REGION Network 63: DeOx/ReOx Valave Configuration Done Sequence Delay
   // Get time value from HMI data
   RUNG wire#powerrail
      Move(in := "86_Times".VLV_CNFG_DN_DLY, out1 => "300_AUT_SEQ_TMRS_DB".VLV_CNFG_DN_DLY.PT)
   END_RUNG
   // the same network as SCL:
   "300_AUT_SEQ_TMRS_DB".VLV_CNFG_DN_DLY.PT := "86_Times".VLV_CNFG_DN_DLY;
END_REGION

REGION Network 64: Modify Maximum Step Time
   // To avoid time-out errors when value changed
   RUNG wire#powerrail
      Add(in1 := "300_AUT_SEQ_TMRS_DB".VLV_CNFG_DN_DLY.PT, in2 := T#100ms, out => "100_GCU_AUTO_SEQ_DB".STEP_410.MST)
   END_RUNG
   // the same network as SCL:
   "100_GCU_AUTO_SEQ_DB".STEP_410.MST := "300_AUT_SEQ_TMRS_DB".VLV_CNFG_DN_DLY.PT + T#100ms;
END_REGION

REGION Network 65: DeOx/ReOx Valave Configuration Done Sequence Delay
   // Run timer
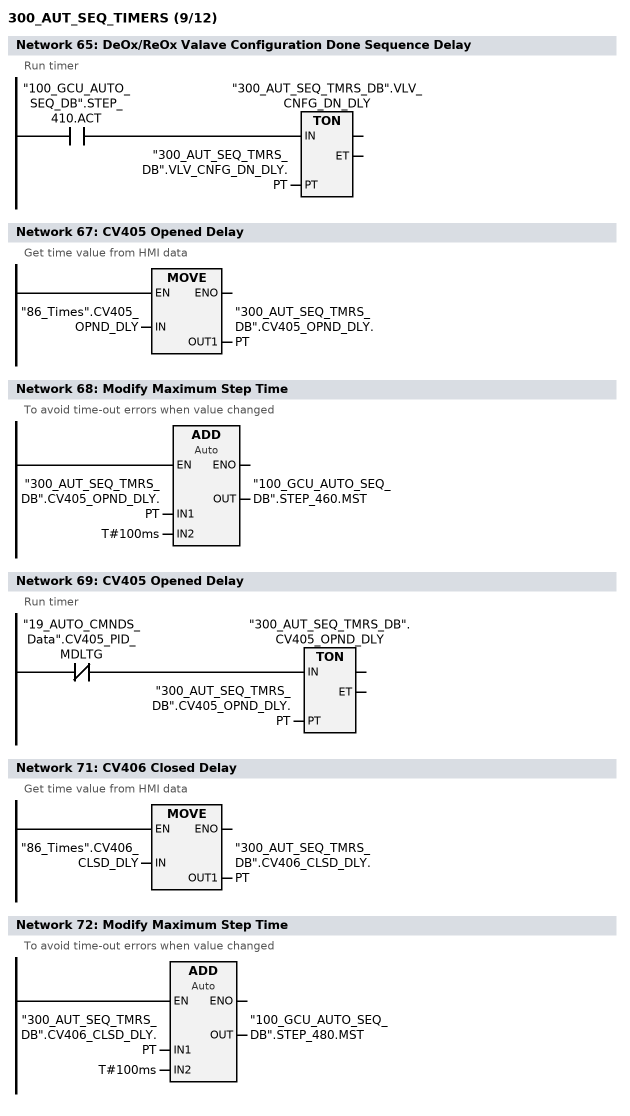
   "300_AUT_SEQ_TMRS_DB".VLV_CNFG_DN_DLY.TON(IN := "100_GCU_AUTO_SEQ_DB".STEP_410.ACT,
                           PT := "300_AUT_SEQ_TMRS_DB".VLV_CNFG_DN_DLY.PT);
END_REGION

REGION Network 67: CV405 Opened Delay
   // Get time value from HMI data
   RUNG wire#powerrail
      Move(in := "86_Times".CV405_OPND_DLY, out1 => "300_AUT_SEQ_TMRS_DB".CV405_OPND_DLY.PT)
   END_RUNG
   // the same network as SCL:
   "300_AUT_SEQ_TMRS_DB".CV405_OPND_DLY.PT := "86_Times".CV405_OPND_DLY;
END_REGION

REGION Network 68: Modify Maximum Step Time
   // To avoid time-out errors when value changed
   RUNG wire#powerrail
      Add(in1 := "300_AUT_SEQ_TMRS_DB".CV405_OPND_DLY.PT, in2 := T#100ms, out => "100_GCU_AUTO_SEQ_DB".STEP_460.MST)
   END_RUNG
   // the same network as SCL:
   "100_GCU_AUTO_SEQ_DB".STEP_460.MST := "300_AUT_SEQ_TMRS_DB".CV405_OPND_DLY.PT + T#100ms;
END_REGION

REGION Network 69: CV405 Opened Delay
   // Run timer
   "300_AUT_SEQ_TMRS_DB".CV405_OPND_DLY.TON(IN := NOT "19_AUTO_CMNDS_Data".CV405_PID_MDLTG,
                           PT := "300_AUT_SEQ_TMRS_DB".CV405_OPND_DLY.PT);
END_REGION

REGION Network 71: CV406 Closed Delay
   // Get time value from HMI data
   RUNG wire#powerrail
      Move(in := "86_Times".CV406_CLSD_DLY, out1 => "300_AUT_SEQ_TMRS_DB".CV406_CLSD_DLY.PT)
   END_RUNG
   // the same network as SCL:
   "300_AUT_SEQ_TMRS_DB".CV406_CLSD_DLY.PT := "86_Times".CV406_CLSD_DLY;
END_REGION

REGION Network 72: Modify Maximum Step Time
   // To avoid time-out errors when value changed
   RUNG wire#powerrail
      Add(in1 := "300_AUT_SEQ_TMRS_DB".CV406_CLSD_DLY.PT, in2 := T#100ms, out => "100_GCU_AUTO_SEQ_DB".STEP_480.MST)
   END_RUNG
   // the same network as SCL:
   "100_GCU_AUTO_SEQ_DB".STEP_480.MST := "300_AUT_SEQ_TMRS_DB".CV406_CLSD_DLY.PT + T#100ms;
END_REGION

REGION Network 73: CV406 Closed Delay
   // Run timer
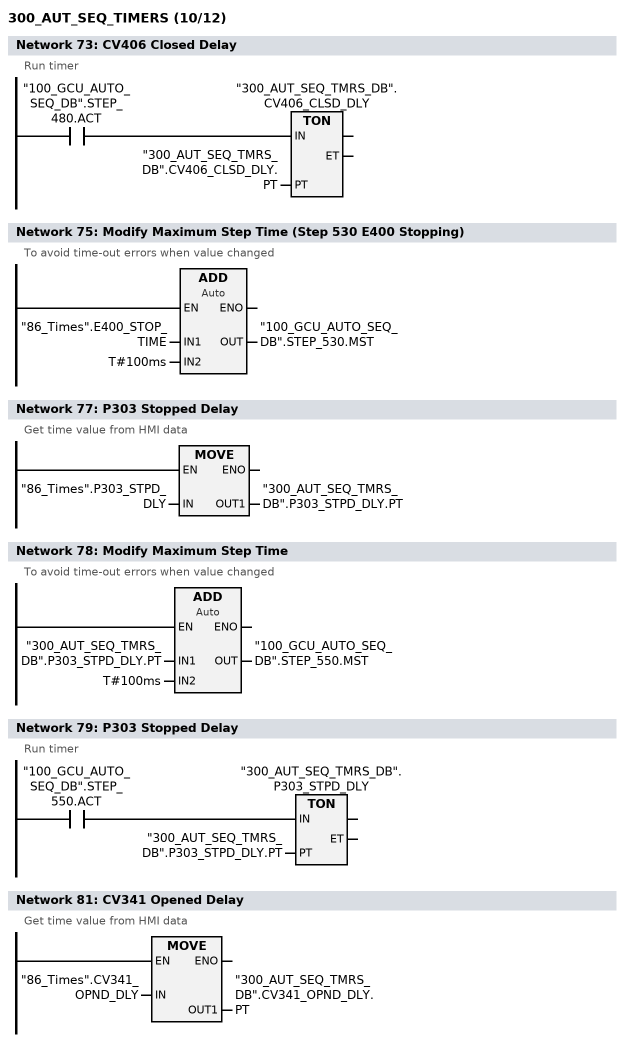
   "300_AUT_SEQ_TMRS_DB".CV406_CLSD_DLY.TON(IN := "100_GCU_AUTO_SEQ_DB".STEP_480.ACT,
                           PT := "300_AUT_SEQ_TMRS_DB".CV406_CLSD_DLY.PT);
END_REGION

REGION Network 75: Modify Maximum Step Time (Step 530 E400 Stopping)
   // To avoid time-out errors when value changed
   RUNG wire#powerrail
      Add(in1 := "86_Times".E400_STOP_TIME, in2 := T#100ms, out => "100_GCU_AUTO_SEQ_DB".STEP_530.MST)
   END_RUNG
   // the same network as SCL:
   "100_GCU_AUTO_SEQ_DB".STEP_530.MST := "86_Times".E400_STOP_TIME + T#100ms;
END_REGION

REGION Network 77: P303 Stopped Delay
   // Get time value from HMI data
   RUNG wire#powerrail
      Move(in := "86_Times".P303_STPD_DLY, out1 => "300_AUT_SEQ_TMRS_DB".P303_STPD_DLY.PT)
   END_RUNG
   // the same network as SCL:
   "300_AUT_SEQ_TMRS_DB".P303_STPD_DLY.PT := "86_Times".P303_STPD_DLY;
END_REGION

REGION Network 78: Modify Maximum Step Time
   // To avoid time-out errors when value changed
   RUNG wire#powerrail
      Add(in1 := "300_AUT_SEQ_TMRS_DB".P303_STPD_DLY.PT, in2 := T#100ms, out => "100_GCU_AUTO_SEQ_DB".STEP_550.MST)
   END_RUNG
   // the same network as SCL:
   "100_GCU_AUTO_SEQ_DB".STEP_550.MST := "300_AUT_SEQ_TMRS_DB".P303_STPD_DLY.PT + T#100ms;
END_REGION

REGION Network 79: P303 Stopped Delay
   // Run timer
   "300_AUT_SEQ_TMRS_DB".P303_STPD_DLY.TON(IN := "100_GCU_AUTO_SEQ_DB".STEP_550.ACT,
                           PT := "300_AUT_SEQ_TMRS_DB".P303_STPD_DLY.PT);
END_REGION

REGION Network 81: CV341 Opened Delay
   // Get time value from HMI data
   RUNG wire#powerrail
      Move(in := "86_Times".CV341_OPND_DLY, out1 => "300_AUT_SEQ_TMRS_DB".CV341_OPND_DLY.PT)
   END_RUNG
   // the same network as SCL:
   "300_AUT_SEQ_TMRS_DB".CV341_OPND_DLY.PT := "86_Times".CV341_OPND_DLY;
END_REGION

REGION Network 82: Modify Maximum Step Time
   // To avoid time-out errors when value changed
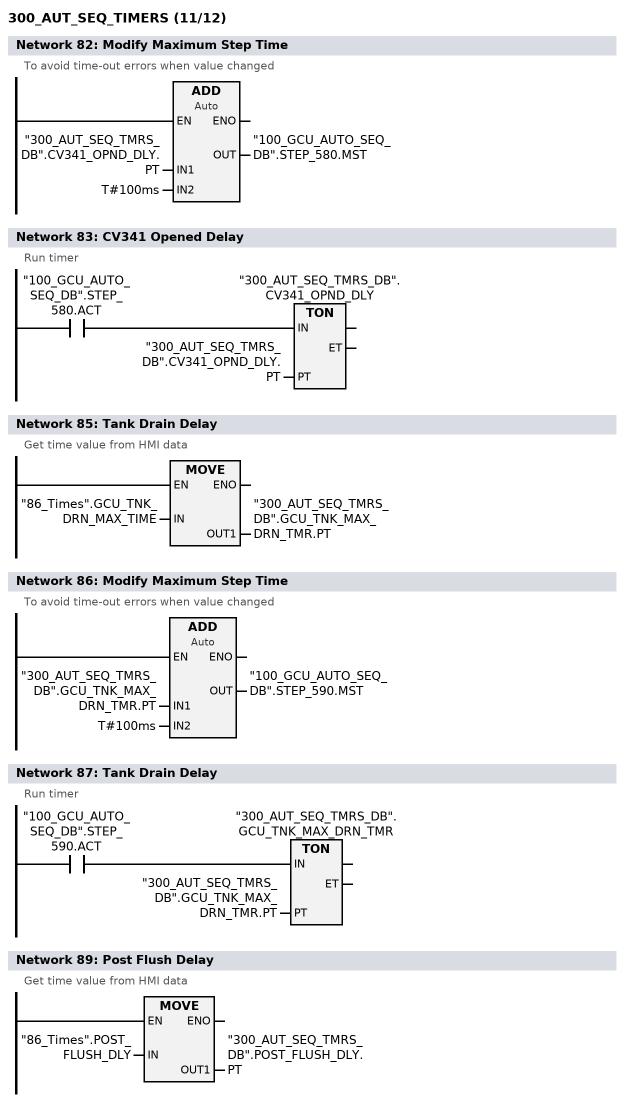
   RUNG wire#powerrail
      Add(in1 := "300_AUT_SEQ_TMRS_DB".CV341_OPND_DLY.PT, in2 := T#100ms, out => "100_GCU_AUTO_SEQ_DB".STEP_580.MST)
   END_RUNG
   // the same network as SCL:
   "100_GCU_AUTO_SEQ_DB".STEP_580.MST := "300_AUT_SEQ_TMRS_DB".CV341_OPND_DLY.PT + T#100ms;
END_REGION

REGION Network 83: CV341 Opened Delay
   // Run timer
   "300_AUT_SEQ_TMRS_DB".CV341_OPND_DLY.TON(IN := "100_GCU_AUTO_SEQ_DB".STEP_580.ACT,
                           PT := "300_AUT_SEQ_TMRS_DB".CV341_OPND_DLY.PT);
END_REGION

REGION Network 85: Tank Drain Delay
   // Get time value from HMI data
   RUNG wire#powerrail
      Move(in := "86_Times".GCU_TNK_DRN_MAX_TIME, out1 => "300_AUT_SEQ_TMRS_DB".GCU_TNK_MAX_DRN_TMR.PT)
   END_RUNG
   // the same network as SCL:
   "300_AUT_SEQ_TMRS_DB".GCU_TNK_MAX_DRN_TMR.PT := "86_Times".GCU_TNK_DRN_MAX_TIME;
END_REGION

REGION Network 86: Modify Maximum Step Time
   // To avoid time-out errors when value changed
   RUNG wire#powerrail
      Add(in1 := "300_AUT_SEQ_TMRS_DB".GCU_TNK_MAX_DRN_TMR.PT, in2 := T#100ms, out => "100_GCU_AUTO_SEQ_DB".STEP_590.MST)
   END_RUNG
   // the same network as SCL:
   "100_GCU_AUTO_SEQ_DB".STEP_590.MST := "300_AUT_SEQ_TMRS_DB".GCU_TNK_MAX_DRN_TMR.PT + T#100ms;
END_REGION

REGION Network 87: Tank Drain Delay
   // Run timer
   "300_AUT_SEQ_TMRS_DB".GCU_TNK_MAX_DRN_TMR.TON(IN := "100_GCU_AUTO_SEQ_DB".STEP_590.ACT,
                           PT := "300_AUT_SEQ_TMRS_DB".GCU_TNK_MAX_DRN_TMR.PT);
END_REGION

REGION Network 89: Post Flush Delay
   // Get time value from HMI data
   RUNG wire#powerrail
      Move(in := "86_Times".POST_FLUSH_DLY, out1 => "300_AUT_SEQ_TMRS_DB".POST_FLUSH_DLY.PT)
   END_RUNG
   // the same network as SCL:
   "300_AUT_SEQ_TMRS_DB".POST_FLUSH_DLY.PT := "86_Times".POST_FLUSH_DLY;
END_REGION

REGION Network 90: Modify Maximum Step Time
   // To avoid time-out errors when value changed
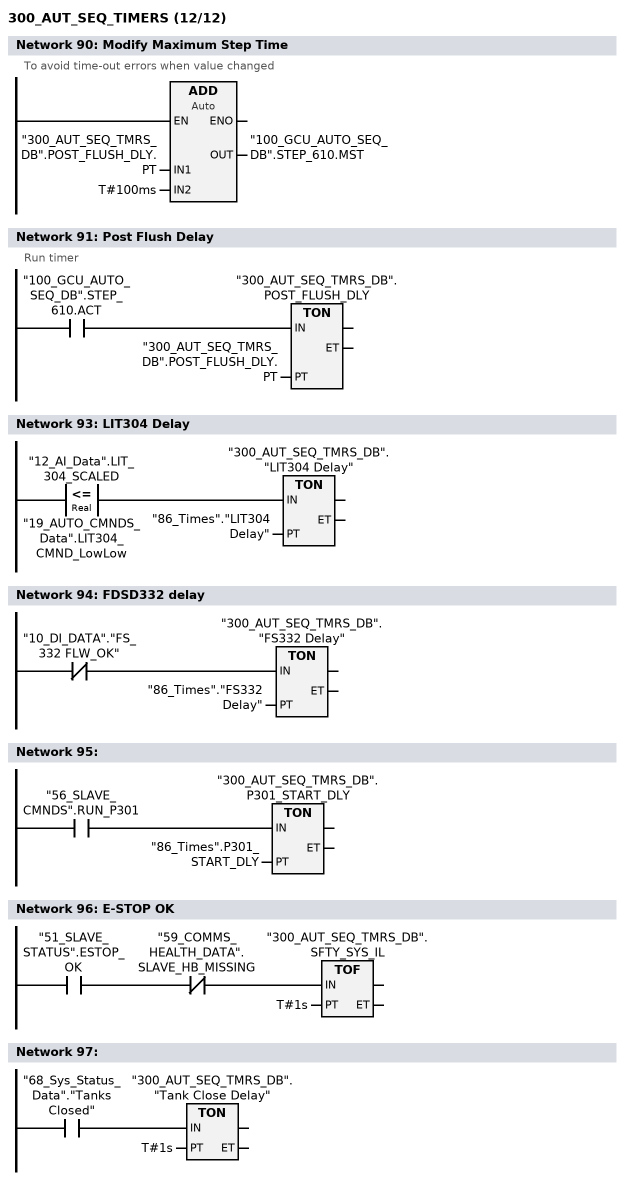
   RUNG wire#powerrail
      Add(in1 := "300_AUT_SEQ_TMRS_DB".POST_FLUSH_DLY.PT, in2 := T#100ms, out => "100_GCU_AUTO_SEQ_DB".STEP_610.MST)
   END_RUNG
   // the same network as SCL:
   "100_GCU_AUTO_SEQ_DB".STEP_610.MST := "300_AUT_SEQ_TMRS_DB".POST_FLUSH_DLY.PT + T#100ms;
END_REGION

REGION Network 91: Post Flush Delay
   // Run timer
   "300_AUT_SEQ_TMRS_DB".POST_FLUSH_DLY.TON(IN := "100_GCU_AUTO_SEQ_DB".STEP_610.ACT,
                           PT := "300_AUT_SEQ_TMRS_DB".POST_FLUSH_DLY.PT);
END_REGION

REGION Network 93: LIT304 Delay
   "300_AUT_SEQ_TMRS_DB"."LIT304 Delay".TON(IN := "12_AI_Data".LIT_304_SCALED <= "19_AUTO_CMNDS_Data".LIT304_CMND_LowLow,
                           PT := "86_Times"."LIT304 Delay");
END_REGION

REGION Network 94: FDSD332 delay
   "300_AUT_SEQ_TMRS_DB"."FS332 Delay".TON(IN := NOT "10_DI_DATA"."FS_332 FLW_OK",
                           PT := "86_Times"."FS332 Delay");
END_REGION

REGION Network 95
   "300_AUT_SEQ_TMRS_DB".P301_START_DLY.TON(IN := "56_SLAVE_CMNDS".RUN_P301, PT := "86_Times".P301_START_DLY);
END_REGION

REGION Network 96: E-STOP OK
   "300_AUT_SEQ_TMRS_DB".SFTY_SYS_IL.TOF(IN := "51_SLAVE_STATUS".ESTOP_OK AND NOT "59_COMMS_HEALTH_DATA".SLAVE_HB_MISSING,
                           PT := T#1s);
END_REGION

REGION Network 97
   "300_AUT_SEQ_TMRS_DB"."Tank Close Delay".TON(IN := "68_Sys_Status_Data"."Tanks Closed", PT := T#1s);
END_REGION
END_FUNCTION

// folder: 50 - 59 PLC Communication

FUNCTION "51_GET_SLAVE_DATA" : Void   // FC51, LAD
TITLE = Get Slave Status Data
{ S7_Optimized_Access := 'TRUE' }
AUTHOR : JRS
VERSION : 0.1
// Code for getting status data from the slave PLC (IGG)
   VAR_TEMP
      RET_VAL_1 : Int;
   END_VAR
BEGIN

REGION Network 1: Get Slave Status Data
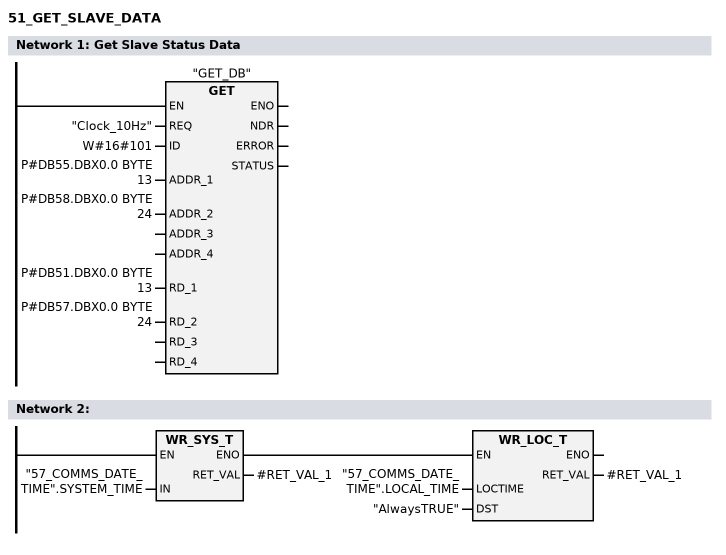
   "GET_DB"(REQ := "Clock_10Hz",   // GET
            ID := W#16#101,
            ADDR_1 := P#DB55.DBX0.0 BYTE 13,
            ADDR_2 := P#DB58.DBX0.0 BYTE 24,
            RD_1 := P#DB51.DBX0.0 BYTE 13,
            RD_2 := P#DB57.DBX0.0 BYTE 24);
END_REGION

REGION Network 2
   // ENO of a box is taken as its EN; it also drops when the box reports an error
   #RET_VAL_1 := WR_SYS_T(IN := "57_COMMS_DATE_TIME".SYSTEM_TIME);
   #RET_VAL_1 := WR_LOC_T(LOCTIME := "57_COMMS_DATE_TIME".LOCAL_TIME, DST := "AlwaysTRUE");
END_REGION
END_FUNCTION

FUNCTION "56_PUT_SLAVE_DATA" : Void   // FC56, LAD
TITLE = Put Slave Comands Data
{ S7_Optimized_Access := 'TRUE' }
AUTHOR : JRS
VERSION : 0.1
// Code for sending commands to the slave PLC (IGG)
BEGIN

REGION Network 1: PUT Slave Commands
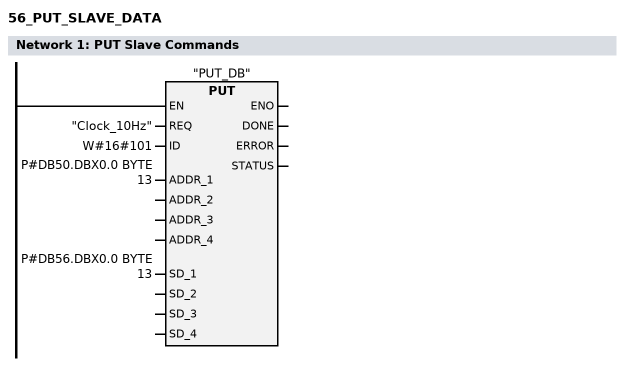
   "PUT_DB"(REQ := "Clock_10Hz", ID := W#16#101, ADDR_1 := P#DB50.DBX0.0 BYTE 13, SD_1 := P#DB56.DBX0.0 BYTE 13);   // PUT
END_REGION
END_FUNCTION

FUNCTION "59_COMMS_HEALTH" : Void   // FC59, LAD
TITLE = Communications Heart Beat
{ S7_Optimized_Access := 'TRUE' }
AUTHOR : JRS
VERSION : 0.1
// Code for communications heart beat bit
   VAR_TEMP   // added for the SCL form of the ladder/FBD networks
      _w1 : Bool;
   END_VAR
BEGIN

REGION Network 1: Local Heart Beat
   // Flip flop for status to other PLC's
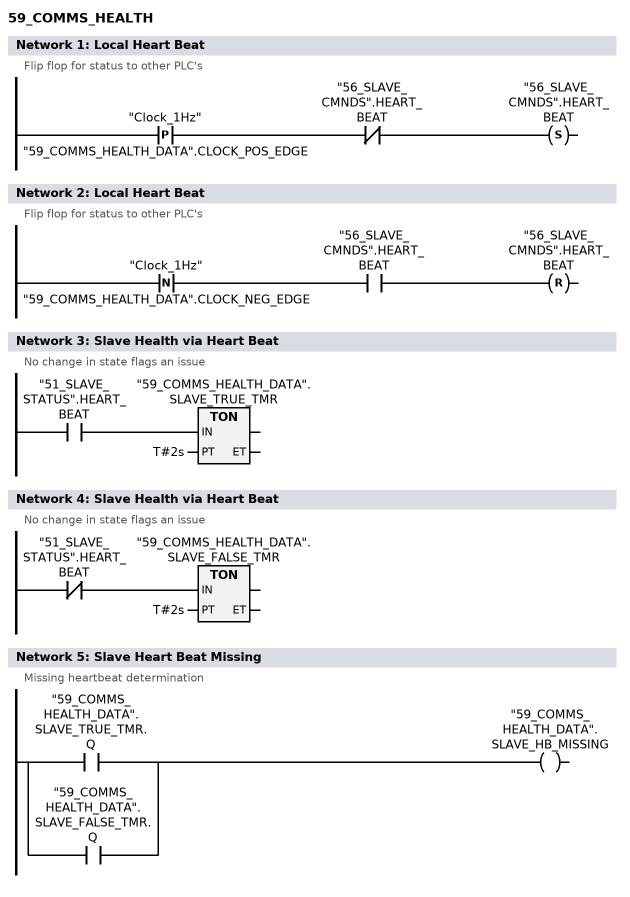
   RUNG wire#powerrail
      P_Contact(operand := "Clock_1Hz", bit := "59_COMMS_HEALTH_DATA".CLOCK_POS_EDGE)
      I_Contact( "56_SLAVE_CMNDS".HEART_BEAT )
      S_Coil( "56_SLAVE_CMNDS".HEART_BEAT )
   END_RUNG
   // the same network as SCL:
   #_w1 := "Clock_1Hz" AND NOT "59_COMMS_HEALTH_DATA".CLOCK_POS_EDGE;   // rising edge of "Clock_1Hz"
   "59_COMMS_HEALTH_DATA".CLOCK_POS_EDGE := "Clock_1Hz";
   IF #_w1 AND NOT "56_SLAVE_CMNDS".HEART_BEAT THEN "56_SLAVE_CMNDS".HEART_BEAT := TRUE; END_IF;
END_REGION

REGION Network 2: Local Heart Beat
   // Flip flop for status to other PLC's
   RUNG wire#powerrail
      N_Contact(operand := "Clock_1Hz", bit := "59_COMMS_HEALTH_DATA".CLOCK_NEG_EDGE)
      Contact( "56_SLAVE_CMNDS".HEART_BEAT )
      R_Coil( "56_SLAVE_CMNDS".HEART_BEAT )
   END_RUNG
   // the same network as SCL:
   #_w1 := NOT "Clock_1Hz" AND "59_COMMS_HEALTH_DATA".CLOCK_NEG_EDGE;   // falling edge of "Clock_1Hz"
   "59_COMMS_HEALTH_DATA".CLOCK_NEG_EDGE := "Clock_1Hz";
   IF #_w1 AND "56_SLAVE_CMNDS".HEART_BEAT THEN "56_SLAVE_CMNDS".HEART_BEAT := FALSE; END_IF;
END_REGION

REGION Network 3: Slave Health via Heart Beat
   // No change in state flags an issue
   "59_COMMS_HEALTH_DATA".SLAVE_TRUE_TMR.TON(IN := "51_SLAVE_STATUS".HEART_BEAT, PT := T#2s);
END_REGION

REGION Network 4: Slave Health via Heart Beat
   // No change in state flags an issue
   "59_COMMS_HEALTH_DATA".SLAVE_FALSE_TMR.TON(IN := NOT "51_SLAVE_STATUS".HEART_BEAT, PT := T#2s);
END_REGION

REGION Network 5: Slave Heart Beat Missing
   // Missing heartbeat determination
   RUNG wire#powerrail
      Contact( "59_COMMS_HEALTH_DATA".SLAVE_TRUE_TMR.Q )
      wire#w1
      Coil( "59_COMMS_HEALTH_DATA".SLAVE_HB_MISSING )
   END_RUNG
   RUNG wire#powerrail
      Contact( "59_COMMS_HEALTH_DATA".SLAVE_FALSE_TMR.Q )
   END_RUNG wire#w1
   // the same network as SCL:
   "59_COMMS_HEALTH_DATA".SLAVE_HB_MISSING := "59_COMMS_HEALTH_DATA".SLAVE_TRUE_TMR.Q OR "59_COMMS_HEALTH_DATA".SLAVE_FALSE_TMR.Q;
END_REGION
END_FUNCTION

// folder: 500 - 699 Standard FBs

FUNCTION_BLOCK "500_SEQ_STEP"   // FB500, LAD
{ S7_Optimized_Access := 'TRUE' }
VERSION : 0.1
   VAR_INPUT
      SN : Int;   // Step number
      CS : Int;   // Current step
      MST : Time;   // Maximum step time
      SC : Bool;   // Step complete
      BPFLT : Bool;   // Bypass fault
   END_VAR
   VAR_OUTPUT
      ACT : Bool;   // Active
      DN : Bool;   // Done
   END_VAR
   VAR_IN_OUT
      AMST : Time;   // Actual maximum step time
      FLT : Bool;   // Timed out
   END_VAR
   VAR
      RNG : Bool;   // Running
   END_VAR
   VAR RETAIN
      STP_MAX_TIM : TON_TIME;   // Maximum step time
   END_VAR
   VAR
      IEC_Timer_0_Instance : TOF_TIME;
   END_VAR
BEGIN

REGION Network 1: Step Active
   // When step number is active, it is also running
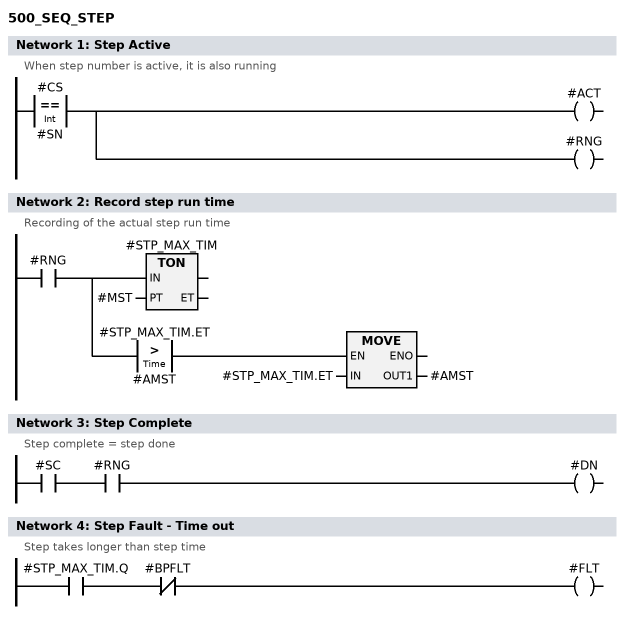
   RUNG wire#powerrail
      { S7_Templates := "SrcType := Int" } EQ_Contact(in1 := #CS, in2 := #SN)
      wire#w1
      Coil( #ACT )
   END_RUNG
   RUNG wire#w1
      Coil( #RNG )
   END_RUNG
   // the same network as SCL:
   #ACT := #CS = #SN;
   #RNG := #ACT;
END_REGION

REGION Network 2: Record step run time
   // Recording of the actual step run time
   #STP_MAX_TIM(IN := #RNG, PT := #MST);   // TON
   IF #RNG AND (#STP_MAX_TIM.ET > #AMST) THEN #AMST := #STP_MAX_TIM.ET; END_IF;
END_REGION

REGION Network 3: Step Complete
   // Step complete = step done
   RUNG wire#powerrail
      Contact( #SC )
      Contact( #RNG )
      Coil( #DN )
   END_RUNG
   // the same network as SCL:
   #DN := #SC AND #RNG;
END_REGION

REGION Network 4: Step Fault - Time out
   // Step takes longer than step time
   RUNG wire#powerrail
      Contact( #STP_MAX_TIM.Q )
      I_Contact( #BPFLT )
      Coil( #FLT )
   END_RUNG
   // the same network as SCL:
   #FLT := #STP_MAX_TIM.Q AND NOT #BPFLT;
END_REGION
END_FUNCTION_BLOCK

FUNCTION_BLOCK "501_VLV_CHK"   // FB501, LAD
TITLE = Valve Check
{ S7_Optimized_Access := 'TRUE' }
AUTHOR : JRS
VERSION : 0.1
// To check for the correct operation of a vlave
   VAR_INPUT
      DMND : Bool;   // Demand
      NO_TYPE : Bool;   // Valve type = open without demand
      NC_TYPE : Bool;   // Valve type = closed without demand
      MAX_MOV_TIM : Time := T#1s;   // Maximum movement time
      OPN_SNSR : Bool;   // Valve open confirmed
      CLS_SNSR : Bool;   // Valve closed confirmed
   END_VAR
   VAR_OUTPUT
      HELTHY : Bool;   // Valve is healthy
      FAULT : Bool;   // Valve is faulty
      CNFG_ERR : Bool;   // Configuration error
   END_VAR
   VAR
      IDLE_FLT : Bool;   // No demand fault
      DMND_FLT : Bool;   // Demand fault
      TRVL_TIME_FLT : Bool;   // Both sensors missing
      SNSR_FLT : Bool;   // Sensor conflicts
      TRVL_TIME : TON_TIME;   // Travel timer
   END_VAR
   // TRVL_TIME.PT := T#1s;
BEGIN

REGION Network 1: Idle Fault
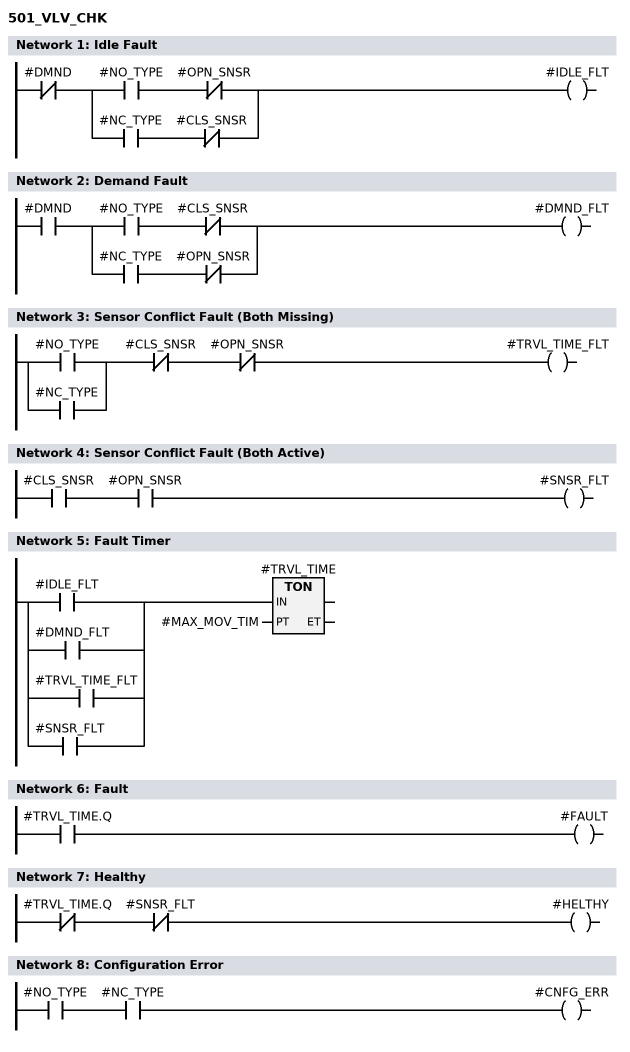
   RUNG wire#powerrail
      I_Contact( #DMND )
      wire#w1
      Contact( #NO_TYPE )
      I_Contact( #OPN_SNSR )
      wire#w2
      Coil( #IDLE_FLT )
   END_RUNG
   RUNG wire#w1
      Contact( #NC_TYPE )
      I_Contact( #CLS_SNSR )
   END_RUNG wire#w2
   // the same network as SCL:
   #IDLE_FLT := NOT #DMND AND ((#NO_TYPE AND NOT #OPN_SNSR) OR (#NC_TYPE AND NOT #CLS_SNSR));
END_REGION

REGION Network 2: Demand Fault
   RUNG wire#powerrail
      Contact( #DMND )
      wire#w1
      Contact( #NO_TYPE )
      I_Contact( #CLS_SNSR )
      wire#w2
      Coil( #DMND_FLT )
   END_RUNG
   RUNG wire#w1
      Contact( #NC_TYPE )
      I_Contact( #OPN_SNSR )
   END_RUNG wire#w2
   // the same network as SCL:
   #DMND_FLT := #DMND AND ((#NO_TYPE AND NOT #CLS_SNSR) OR (#NC_TYPE AND NOT #OPN_SNSR));
END_REGION

REGION Network 3: Sensor Conflict Fault (Both Missing)
   RUNG wire#powerrail
      Contact( #NO_TYPE )
      wire#w1
      I_Contact( #CLS_SNSR )
      I_Contact( #OPN_SNSR )
      Coil( #TRVL_TIME_FLT )
   END_RUNG
   RUNG wire#powerrail
      Contact( #NC_TYPE )
   END_RUNG wire#w1
   // the same network as SCL:
   #TRVL_TIME_FLT := (#NO_TYPE OR #NC_TYPE) AND NOT #CLS_SNSR AND NOT #OPN_SNSR;
END_REGION

REGION Network 4: Sensor Conflict Fault (Both Active)
   RUNG wire#powerrail
      Contact( #CLS_SNSR )
      Contact( #OPN_SNSR )
      Coil( #SNSR_FLT )
   END_RUNG
   // the same network as SCL:
   #SNSR_FLT := #CLS_SNSR AND #OPN_SNSR;
END_REGION

REGION Network 5: Fault Timer
   #TRVL_TIME(IN := #IDLE_FLT OR #DMND_FLT OR #TRVL_TIME_FLT OR #SNSR_FLT, PT := #MAX_MOV_TIM);   // TON
END_REGION

REGION Network 6: Fault
   RUNG wire#powerrail
      Contact( #TRVL_TIME.Q )
      Coil( #FAULT )
   END_RUNG
   // the same network as SCL:
   #FAULT := #TRVL_TIME.Q;
END_REGION

REGION Network 7: Healthy
   RUNG wire#powerrail
      I_Contact( #TRVL_TIME.Q )
      I_Contact( #SNSR_FLT )
      Coil( #HELTHY )
   END_RUNG
   // the same network as SCL:
   #HELTHY := NOT #TRVL_TIME.Q AND NOT #SNSR_FLT;
END_REGION

REGION Network 8: Configuration Error
   RUNG wire#powerrail
      Contact( #NO_TYPE )
      Contact( #NC_TYPE )
      Coil( #CNFG_ERR )
   END_RUNG
   // the same network as SCL:
   #CNFG_ERR := #NO_TYPE AND #NC_TYPE;
END_REGION
END_FUNCTION_BLOCK

FUNCTION_BLOCK "502_ALM_ANALOG"   // FB502, LAD
{ S7_Optimized_Access := 'FALSE' }
VERSION : 0.1
   VAR_INPUT
      Value : Real;
      "Raw Value" : Int;
      Enable : Bool := true;
      "Enable Delay Time" : Time := T#10s;
      "High Value Release" : Bool := true;   // It is Releasing High Values from Enable restriction
      "SHORT CIRCUIT VALUE" : Real := 32000.0;
      "BROKEN WIRE VALUE" : Real := -32000.0;
      "VERY LOW LEVEL VALUE (LL)" : Real;
      "LOW LEVEL VALUE (L)" : Real;
      "HIGH LEVEL VALUE (H)" : Real;
      "VERY HIGH LEVEL VALUE (HH)" : Real;
      OFFSET : Real;
      "ALARM DELAY" : Time := T#1s;
      "Peak Value Reset" : Bool;
   END_VAR
   VAR_OUTPUT
      "ALARM HH" : Bool;
      "ALARM H" : Bool;
      "ALARM L" : Bool;
      "ALARM LL" : Bool;
      "ALARM READING" : Bool;
      "Peak Value" : Real;
      Alarm : Word;
      Alarm_INT : Int;
   END_VAR
   VAR
      TRUE : Bool;
      FALSE : Bool;
      Raw_value_int : Int;
      RET_VAL : Word;
      RAW_scaled_mA : Real;
      RAW_scaled_VALUE : Real;
      SCALED_OFFSETTED_VALUE : Real;
      Error_present : Bool;
      "Enable Internal" : Bool;
      "ALARM HH_interm" : Bool;
      "ALARM H_interm" : Bool;
      "ALARM L_interm" : Bool;
      "ALARM LL_interm" : Bool;
      "ALARM READING_interm" : Bool;
      "ALARM_HH delay" : TON_TIME;
      "ALARM_H delay" : TON_TIME;
      "ALARM_LL delay" : TON_TIME;
      "ALARM_L delay" : TON_TIME;
      "ALARM_READING delay" : TON_TIME;
      "ALARM READING TOF" : TOF_TIME;
      "HI HI TOF" : TOF_TIME;
      "HI TOF" : TOF_TIME;
      "LOE TOF" : TOF_TIME;
      "LOW TOF" : TOF_TIME;
      "LOW LOW TOF" : TOF_TIME;
      "Enable TON" : TON_TIME;
   END_VAR
   VAR_TEMP   // added for the SCL form of the ladder/FBD networks
      _w1 : Bool;
   END_VAR
BEGIN

REGION Network 1: True False
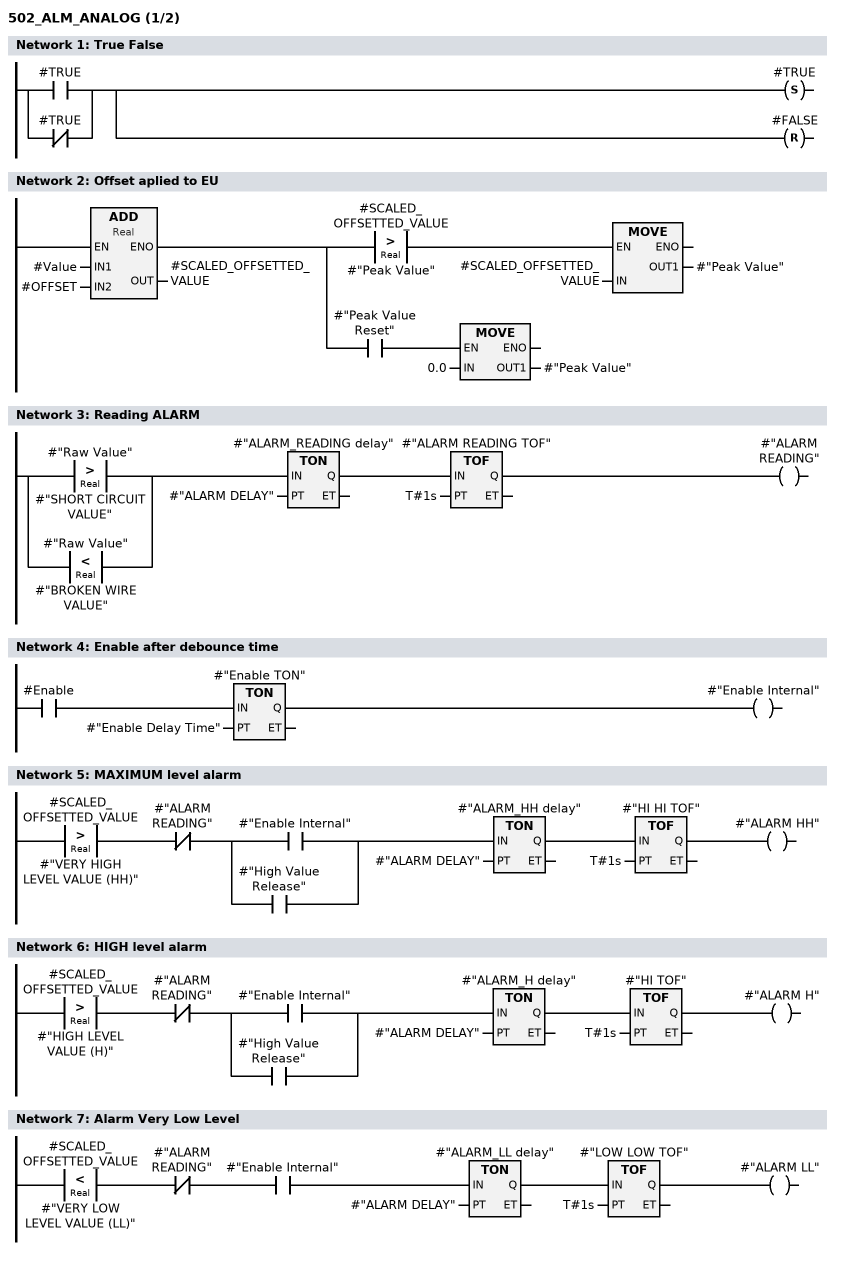
   RUNG wire#powerrail
      Contact( #TRUE )
      wire#w1
      S_Coil( #TRUE )
   END_RUNG
   RUNG wire#powerrail
      I_Contact( #TRUE )
   END_RUNG wire#w1
   RUNG wire#w1
      R_Coil( #FALSE )
   END_RUNG
   // the same network as SCL:
   #_w1 := #TRUE OR NOT #TRUE;
   IF #_w1 THEN
       #TRUE := TRUE;
       #FALSE := FALSE;
   END_IF;
END_REGION

REGION Network 2: Offset aplied to EU
   RUNG wire#powerrail
      { S7_Templates := "SrcType := Real"; S7_GenerateENO := "TRUE" } Add(in1 := #Value, in2 := #OFFSET, out => #SCALED_OFFSETTED_VALUE)
      wire#w1
      { S7_Templates := "SrcType := Real" } GT_Contact(in1 := #SCALED_OFFSETTED_VALUE, in2 := #"Peak Value")
      Move(in := #SCALED_OFFSETTED_VALUE, out1 => #"Peak Value")
   END_RUNG
   RUNG wire#w1
      Contact( #"Peak Value Reset" )
      Move(in := 0.0, out1 => #"Peak Value")
   END_RUNG
   // the same network as SCL:
   // ENO of a box is taken as its EN; it also drops when the box reports an error
   #SCALED_OFFSETTED_VALUE := #Value + #OFFSET;
   IF #SCALED_OFFSETTED_VALUE > #"Peak Value" THEN #"Peak Value" := #SCALED_OFFSETTED_VALUE; END_IF;
   IF #"Peak Value Reset" THEN #"Peak Value" := 0.0; END_IF;
END_REGION

REGION Network 3: Reading ALARM
   #"ALARM_READING delay"(IN := (#"Raw Value" > #"SHORT CIRCUIT VALUE") OR (#"Raw Value" < #"BROKEN WIRE VALUE"),   // TON
                          PT := #"ALARM DELAY");
   #"ALARM READING TOF"(IN := #"ALARM_READING delay".Q, PT := T#1s);   // TOF
   #"ALARM READING" := #"ALARM READING TOF".Q;
END_REGION

REGION Network 4: Enable after debounce time
   #"Enable TON"(IN := #Enable, PT := #"Enable Delay Time");   // TON
   #"Enable Internal" := #"Enable TON".Q;
END_REGION

REGION Network 5: MAXIMUM level alarm
   #"ALARM_HH delay"(IN := (#SCALED_OFFSETTED_VALUE > #"VERY HIGH LEVEL VALUE (HH)") AND NOT #"ALARM READING" AND (#"Enable Internal" OR #"High Value Release"),   // TON
                     PT := #"ALARM DELAY");
   #"HI HI TOF"(IN := #"ALARM_HH delay".Q, PT := T#1s);   // TOF
   #"ALARM HH" := #"HI HI TOF".Q;
END_REGION

REGION Network 6: HIGH level alarm
   #"ALARM_H delay"(IN := (#SCALED_OFFSETTED_VALUE > #"HIGH LEVEL VALUE (H)") AND NOT #"ALARM READING" AND (#"Enable Internal" OR #"High Value Release"),   // TON
                    PT := #"ALARM DELAY");
   #"HI TOF"(IN := #"ALARM_H delay".Q, PT := T#1s);   // TOF
   #"ALARM H" := #"HI TOF".Q;
END_REGION

REGION Network 7: Alarm Very Low Level
   #"ALARM_LL delay"(IN := (#SCALED_OFFSETTED_VALUE < #"VERY LOW LEVEL VALUE (LL)") AND NOT #"ALARM READING" AND #"Enable Internal",   // TON
                     PT := #"ALARM DELAY");
   #"LOW LOW TOF"(IN := #"ALARM_LL delay".Q, PT := T#1s);   // TOF
   #"ALARM LL" := #"LOW LOW TOF".Q;
END_REGION

REGION Network 8: Alarm Low Level
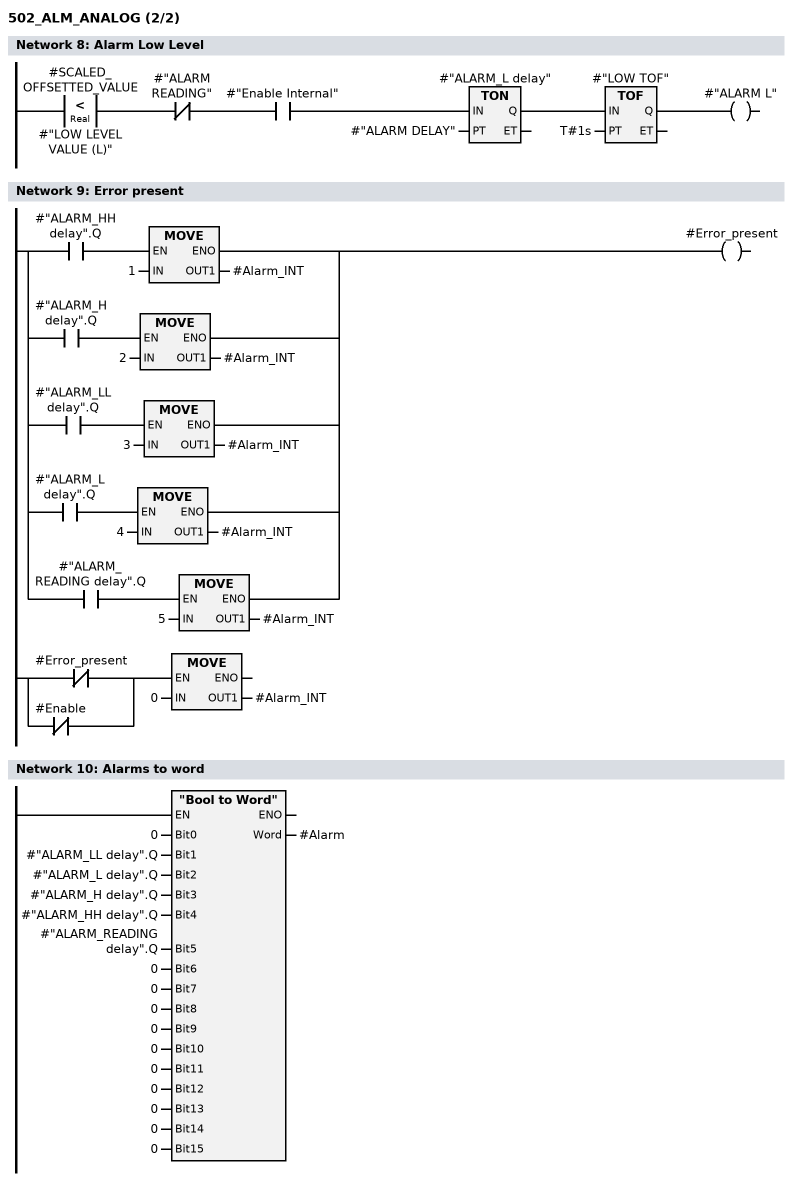
   #"ALARM_L delay"(IN := (#SCALED_OFFSETTED_VALUE < #"LOW LEVEL VALUE (L)") AND NOT #"ALARM READING" AND #"Enable Internal",   // TON
                    PT := #"ALARM DELAY");
   #"LOW TOF"(IN := #"ALARM_L delay".Q, PT := T#1s);   // TOF
   #"ALARM L" := #"LOW TOF".Q;
END_REGION

REGION Network 9: Error present
   RUNG wire#powerrail
      Contact( #"ALARM_HH delay".Q )
      { S7_GenerateENO := "TRUE" } Move(in := 1, out1 => #Alarm_INT)
      wire#w1
      Coil( #Error_present )
   END_RUNG
   RUNG wire#powerrail
      Contact( #"ALARM_H delay".Q )
      { S7_GenerateENO := "TRUE" } Move(in := 2, out1 => #Alarm_INT)
   END_RUNG wire#w1
   RUNG wire#powerrail
      Contact( #"ALARM_LL delay".Q )
      { S7_GenerateENO := "TRUE" } Move(in := 3, out1 => #Alarm_INT)
   END_RUNG wire#w1
   RUNG wire#powerrail
      Contact( #"ALARM_L delay".Q )
      { S7_GenerateENO := "TRUE" } Move(in := 4, out1 => #Alarm_INT)
   END_RUNG wire#w1
   RUNG wire#powerrail
      Contact( #"ALARM_READING delay".Q )
      { S7_GenerateENO := "TRUE" } Move(in := 5, out1 => #Alarm_INT)
   END_RUNG wire#w1
   RUNG wire#powerrail
      I_Contact( #Error_present )
      wire#w2
      Move(in := 0, out1 => #Alarm_INT)
   END_RUNG
   RUNG wire#powerrail
      I_Contact( #Enable )
   END_RUNG wire#w2
   // the same network as SCL:
   // ENO of a box is taken as its EN; it also drops when the box reports an error
   IF #"ALARM_HH delay".Q THEN #Alarm_INT := 1; END_IF;
   IF #"ALARM_H delay".Q THEN #Alarm_INT := 2; END_IF;
   IF #"ALARM_LL delay".Q THEN #Alarm_INT := 3; END_IF;
   IF #"ALARM_L delay".Q THEN #Alarm_INT := 4; END_IF;
   IF #"ALARM_READING delay".Q THEN #Alarm_INT := 5; END_IF;
   #Error_present := #"ALARM_HH delay".Q OR #"ALARM_H delay".Q OR #"ALARM_LL delay".Q OR #"ALARM_L delay".Q OR #"ALARM_READING delay".Q;
   IF NOT #Error_present OR NOT #Enable THEN #Alarm_INT := 0; END_IF;
END_REGION

REGION Network 10: Alarms to word
   RUNG wire#powerrail
      "Bool to Word"(Bit0 := 0, Bit1 := #"ALARM_LL delay".Q, Bit2 := #"ALARM_L delay".Q, Bit3 := #"ALARM_H delay".Q, Bit4 := #"ALARM_HH delay".Q, Bit5 := #"ALARM_READING delay".Q, Bit6 := 0, Bit7 := 0, Bit8 := 0, Bit9 := 0, Bit10 := 0, Bit11 := 0, Bit12 := 0, Bit13 := 0, Bit14 := 0, Bit15 := 0, "Word" => #Alarm)
   END_RUNG
   // the same network as SCL:
   "Bool to Word"(Bit0 := 0,
                  Bit1 := #"ALARM_LL delay".Q,
                  Bit2 := #"ALARM_L delay".Q,
                  Bit3 := #"ALARM_H delay".Q,
                  Bit4 := #"ALARM_HH delay".Q,
                  Bit5 := #"ALARM_READING delay".Q,
                  Bit6 := 0,
                  Bit7 := 0,
                  Bit8 := 0,
                  Bit9 := 0,
                  Bit10 := 0,
                  Bit11 := 0,
                  Bit12 := 0,
                  Bit13 := 0,
                  Bit14 := 0,
                  Bit15 := 0,
                  "Word" => #Alarm);
END_REGION
END_FUNCTION_BLOCK

FUNCTION_BLOCK "Tank Grouping"   // FB504, LAD
TITLE = Tank Grouping
{ S7_Optimized_Access := 'TRUE' }
AUTHOR : Adrian_Stefanescu